REGION Network 21: FC_CARGA_RECETA
   RUNG wire#powerrail
      Contact( "flanco"."pHMI.Pls_CargarReceta" )
      "FC_CARGA_RECETA"("NRO RECETA" := "DB_Animación".Nro_Receta_Edición)
   END_RUNG
   // the same network as SCL:
   IF "flanco"."pHMI.Pls_CargarReceta" THEN
       "FC_CARGA_RECETA"("NRO RECETA" := "DB_Animación".Nro_Receta_Edición);
   END_IF;
END_REGION

REGION Network 22: Proceso a Animación
   RUNG wire#powerrail
      I_Contact( "Editando_Recetas" )
      "CAPA Proceso_Animación"()
   END_RUNG
   // the same network as SCL:
   IF NOT "Editando_Recetas" THEN "CAPA Proceso_Animación"(); END_IF;
END_REGION

REGION Network 23: CAPA Receta_Animación_Receta
   RUNG wire#powerrail
      "CAPA Receta_Animación_Receta"()
   END_RUNG
   // the same network as SCL:
   "CAPA Receta_Animación_Receta"();
END_REGION

REGION Network 24: Animación
   RUNG wire#powerrail
      "FC_Animación"()
   END_RUNG
   // the same network as SCL:
   "FC_Animación"();
END_REGION

REGION Network 25: RESET ELEM ACTUAL
   RUNG wire#powerrail
      I_Contact( "AUTO/MAN" )
      "FC_RESET_ELEM_ACTUAL"()
   END_RUNG
   // the same network as SCL:
   IF NOT "AUTO/MAN" THEN "FC_RESET_ELEM_ACTUAL"(); END_IF;
END_REGION

REGION Network 26: Alarmas
   RUNG wire#powerrail
      "10_FC_Alarmas"()
   END_RUNG
   // the same network as SCL:
   "10_FC_Alarmas"();
END_REGION

REGION Network 27: Salidas
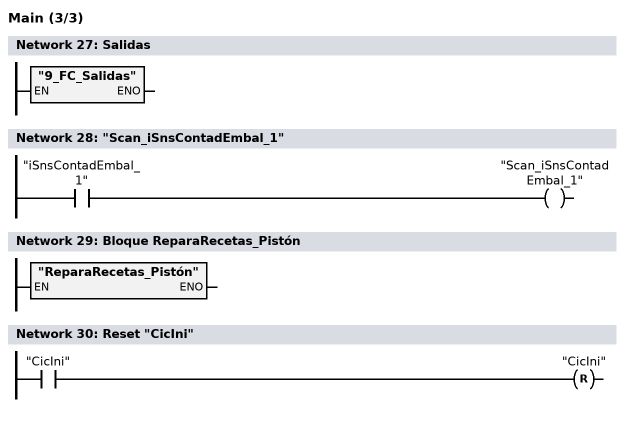
   RUNG wire#powerrail
      "9_FC_Salidas"()
   END_RUNG
   // the same network as SCL:
   "9_FC_Salidas"();
END_REGION

REGION Network 28: "Scan_iSnsContadEmbal_1"
   RUNG wire#powerrail
      Contact( "iSnsContadEmbal_1" )
      Coil( "Scan_iSnsContadEmbal_1" )
   END_RUNG
   // the same network as SCL:
   "Scan_iSnsContadEmbal_1" := "iSnsContadEmbal_1";
END_REGION

REGION Network 29: Bloque ReparaRecetas_Pistón
   RUNG wire#powerrail
      "ReparaRecetas_Pistón"()
   END_RUNG
   // the same network as SCL:
   "ReparaRecetas_Pistón"();
END_REGION

REGION Network 30: Reset "CicIni"
   RUNG wire#powerrail
      Contact( "CicIni" )
      R_Coil( "CicIni" )
   END_RUNG
   // the same network as SCL:
   IF "CicIni" THEN "CicIni" := FALSE; END_IF;
END_REGION
END_ORGANIZATION_BLOCK

ORGANIZATION_BLOCK "CYCL_FLT"   // OB80, LAD
TITLE = "Cycle Time Fault"
{ S7_Optimized_Access := 'FALSE' }
VERSION : 0.1
BEGIN
END_ORGANIZATION_BLOCK

ORGANIZATION_BLOCK "I/O_FLT1"   // OB82, LAD
TITLE = "I/O Point Fault"
{ S7_Optimized_Access := 'FALSE' }
VERSION : 0.1
BEGIN
END_ORGANIZATION_BLOCK

ORGANIZATION_BLOCK "OBNL_FLT"   // OB85, LAD
TITLE = "Organization Block (OB) Not Loaded Fault"
{ S7_Optimized_Access := 'FALSE' }
VERSION : 0.1
BEGIN
END_ORGANIZATION_BLOCK

ORGANIZATION_BLOCK "COMM_FLT"   // OB87, LAD
TITLE = "Communication Fault"
{ S7_Optimized_Access := 'FALSE' }
VERSION : 0.1
BEGIN
END_ORGANIZATION_BLOCK

ORGANIZATION_BLOCK "COMPLETE RESTART"   // OB100, LAD
TITLE = "Complete Restart"
{ S7_Optimized_Access := 'FALSE' }
VERSION : 0.1
BEGIN

REGION Network 1: "bit1"
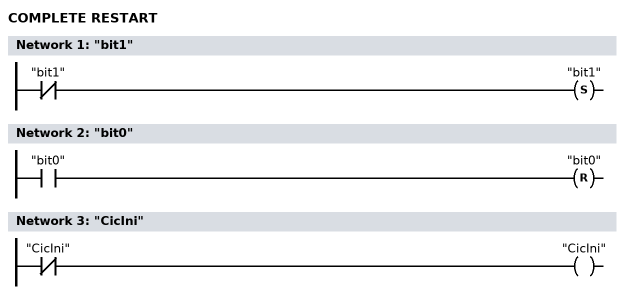
   RUNG wire#powerrail
      I_Contact( "bit1" )
      S_Coil( "bit1" )
   END_RUNG
   // the same network as SCL:
   IF NOT "bit1" THEN "bit1" := TRUE; END_IF;
END_REGION

REGION Network 2: "bit0"
   RUNG wire#powerrail
      Contact( "bit0" )
      R_Coil( "bit0" )
   END_RUNG
   // the same network as SCL:
   IF "bit0" THEN "bit0" := FALSE; END_IF;
END_REGION

REGION Network 3: "CicIni"
   RUNG wire#powerrail
      I_Contact( "CicIni" )
      Coil( "CicIni" )
   END_RUNG
   // the same network as SCL:
   "CicIni" := NOT "CicIni";
END_REGION
END_ORGANIZATION_BLOCK

ORGANIZATION_BLOCK "PROG_ERR"   // OB121, LAD
TITLE = "Programming Error"
{ S7_Optimized_Access := 'FALSE' }
VERSION : 0.1
BEGIN
END_ORGANIZATION_BLOCK

ORGANIZATION_BLOCK "MOD_ERR"   // OB122, LAD
TITLE = "Module Access Error"
{ S7_Optimized_Access := 'FALSE' }
VERSION : 0.1
BEGIN
END_ORGANIZATION_BLOCK

// folder: Alarmas

FUNCTION "10_FC_Alarmas" : Void   // FC23, LAD
{ S7_Optimized_Access := 'FALSE' }
VERSION : 0.1
BEGIN

REGION Network 1: Falla 1: Emergencia Almacén Pallets
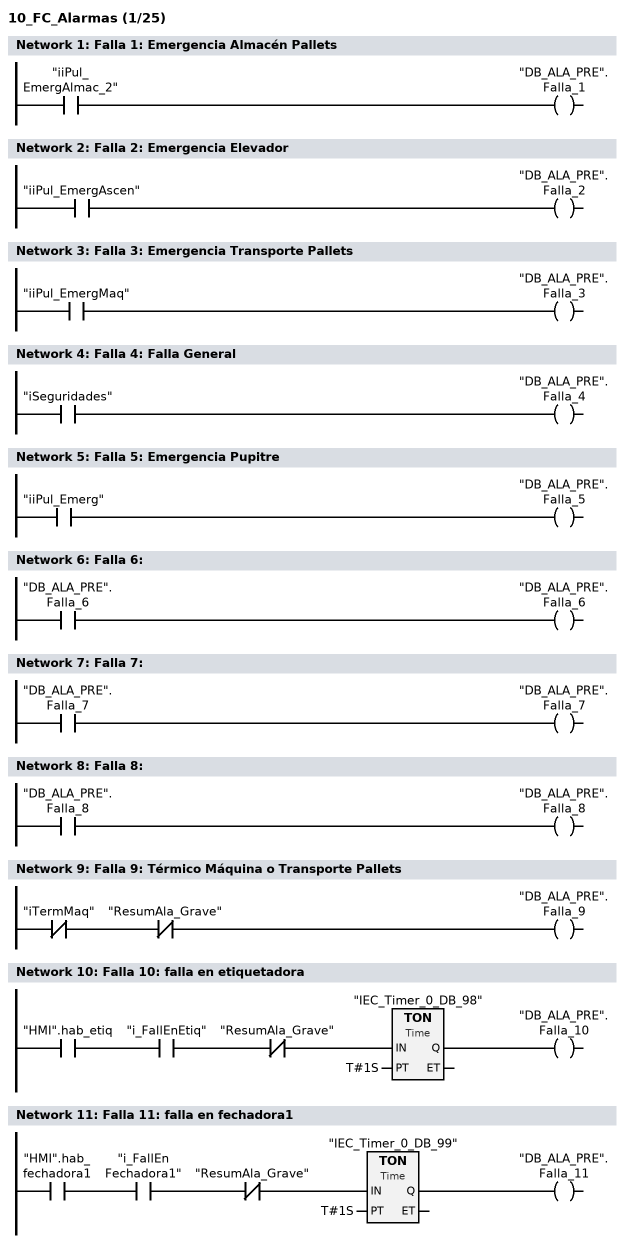
   RUNG wire#powerrail
      Contact( "iiPul_EmergAlmac_2" )
      Coil( "DB_ALA_PRE".Falla_1 )
   END_RUNG
   // the same network as SCL:
   "DB_ALA_PRE".Falla_1 := "iiPul_EmergAlmac_2";
END_REGION

REGION Network 2: Falla 2: Emergencia Elevador
   RUNG wire#powerrail
      Contact( "iiPul_EmergAscen" )
      Coil( "DB_ALA_PRE".Falla_2 )
   END_RUNG
   // the same network as SCL:
   "DB_ALA_PRE".Falla_2 := "iiPul_EmergAscen";
END_REGION

REGION Network 3: Falla 3: Emergencia Transporte Pallets
   RUNG wire#powerrail
      Contact( "iiPul_EmergMaq" )
      Coil( "DB_ALA_PRE".Falla_3 )
   END_RUNG
   // the same network as SCL:
   "DB_ALA_PRE".Falla_3 := "iiPul_EmergMaq";
END_REGION

REGION Network 4: Falla 4: Falla General
   RUNG wire#powerrail
      Contact( "iSeguridades" )
      Coil( "DB_ALA_PRE".Falla_4 )
   END_RUNG
   // the same network as SCL:
   "DB_ALA_PRE".Falla_4 := "iSeguridades";
END_REGION

REGION Network 5: Falla 5: Emergencia Pupitre
   RUNG wire#powerrail
      Contact( "iiPul_Emerg" )
      Coil( "DB_ALA_PRE".Falla_5 )
   END_RUNG
   // the same network as SCL:
   "DB_ALA_PRE".Falla_5 := "iiPul_Emerg";
END_REGION

REGION Network 6: Falla 6:
   RUNG wire#powerrail
      Contact( "DB_ALA_PRE".Falla_6 )
      Coil( "DB_ALA_PRE".Falla_6 )
   END_RUNG
   // the same network as SCL:
   "DB_ALA_PRE".Falla_6 := "DB_ALA_PRE".Falla_6;
END_REGION

REGION Network 7: Falla 7:
   RUNG wire#powerrail
      Contact( "DB_ALA_PRE".Falla_7 )
      Coil( "DB_ALA_PRE".Falla_7 )
   END_RUNG
   // the same network as SCL:
   "DB_ALA_PRE".Falla_7 := "DB_ALA_PRE".Falla_7;
END_REGION

REGION Network 8: Falla 8:
   RUNG wire#powerrail
      Contact( "DB_ALA_PRE".Falla_8 )
      Coil( "DB_ALA_PRE".Falla_8 )
   END_RUNG
   // the same network as SCL:
   "DB_ALA_PRE".Falla_8 := "DB_ALA_PRE".Falla_8;
END_REGION

REGION Network 9: Falla 9: Térmico Máquina o Transporte Pallets
   RUNG wire#powerrail
      I_Contact( "iTermMaq" )
      I_Contact( "ResumAla_Grave" )
      Coil( "DB_ALA_PRE".Falla_9 )
   END_RUNG
   // the same network as SCL:
   "DB_ALA_PRE".Falla_9 := NOT "iTermMaq" AND NOT "ResumAla_Grave";
END_REGION

REGION Network 10: Falla 10: falla en etiquetadora
   "IEC_Timer_0_DB_98".TON(IN := "HMI".hab_etiq AND "i_FallEnEtiq" AND NOT "ResumAla_Grave", PT := T#1S);
   "DB_ALA_PRE".Falla_10 := "IEC_Timer_0_DB_98".Q;
END_REGION

REGION Network 11: Falla 11: falla en fechadora1
   "IEC_Timer_0_DB_99".TON(IN := "HMI".hab_fechadora1 AND "i_FallEnFechadora1" AND NOT "ResumAla_Grave",
                           PT := T#1S);
   "DB_ALA_PRE".Falla_11 := "IEC_Timer_0_DB_99".Q;
END_REGION

REGION Network 12: Falla 12: falla en fechadora2
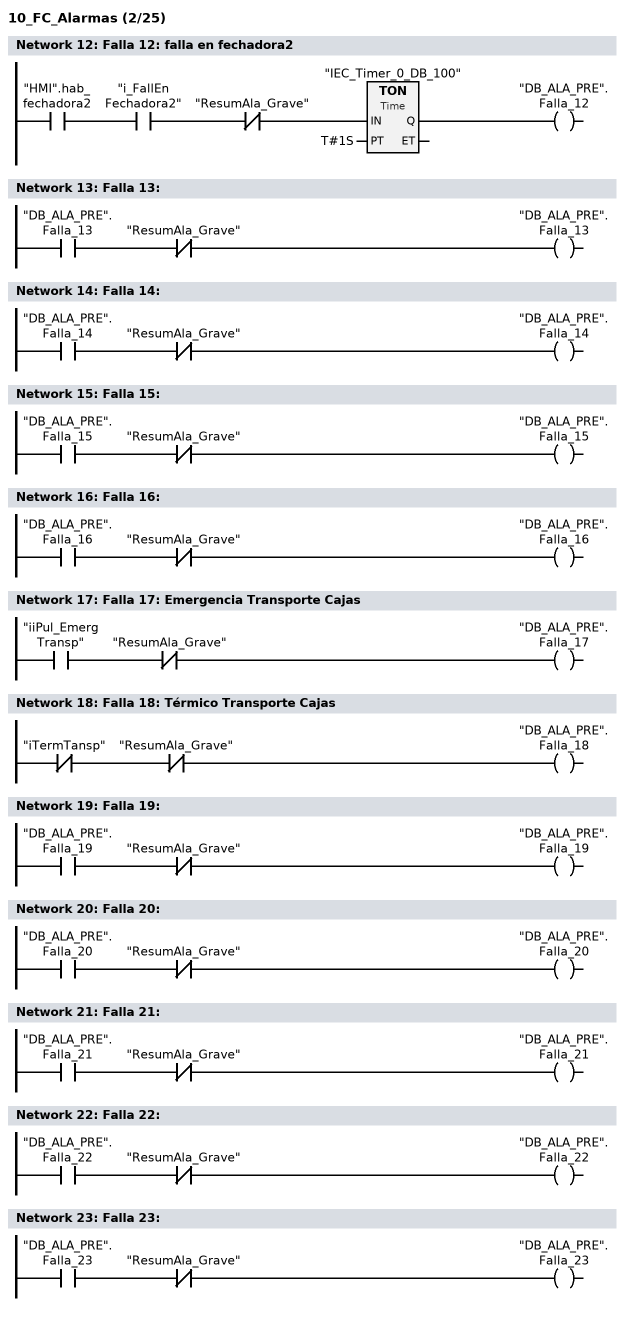
   "IEC_Timer_0_DB_100".TON(IN := "HMI".hab_fechadora2 AND "i_FallEnFechadora2" AND NOT "ResumAla_Grave",
                           PT := T#1S);
   "DB_ALA_PRE".Falla_12 := "IEC_Timer_0_DB_100".Q;
END_REGION

REGION Network 13: Falla 13:
   RUNG wire#powerrail
      Contact( "DB_ALA_PRE".Falla_13 )
      I_Contact( "ResumAla_Grave" )
      Coil( "DB_ALA_PRE".Falla_13 )
   END_RUNG
   // the same network as SCL:
   "DB_ALA_PRE".Falla_13 := "DB_ALA_PRE".Falla_13 AND NOT "ResumAla_Grave";
END_REGION

REGION Network 14: Falla 14:
   RUNG wire#powerrail
      Contact( "DB_ALA_PRE".Falla_14 )
      I_Contact( "ResumAla_Grave" )
      Coil( "DB_ALA_PRE".Falla_14 )
   END_RUNG
   // the same network as SCL:
   "DB_ALA_PRE".Falla_14 := "DB_ALA_PRE".Falla_14 AND NOT "ResumAla_Grave";
END_REGION

REGION Network 15: Falla 15:
   RUNG wire#powerrail
      Contact( "DB_ALA_PRE".Falla_15 )
      I_Contact( "ResumAla_Grave" )
      Coil( "DB_ALA_PRE".Falla_15 )
   END_RUNG
   // the same network as SCL:
   "DB_ALA_PRE".Falla_15 := "DB_ALA_PRE".Falla_15 AND NOT "ResumAla_Grave";
END_REGION

REGION Network 16: Falla 16:
   RUNG wire#powerrail
      Contact( "DB_ALA_PRE".Falla_16 )
      I_Contact( "ResumAla_Grave" )
      Coil( "DB_ALA_PRE".Falla_16 )
   END_RUNG
   // the same network as SCL:
   "DB_ALA_PRE".Falla_16 := "DB_ALA_PRE".Falla_16 AND NOT "ResumAla_Grave";
END_REGION

REGION Network 17: Falla 17: Emergencia Transporte Cajas
   RUNG wire#powerrail
      Contact( "iiPul_EmergTransp" )
      I_Contact( "ResumAla_Grave" )
      Coil( "DB_ALA_PRE".Falla_17 )
   END_RUNG
   // the same network as SCL:
   "DB_ALA_PRE".Falla_17 := "iiPul_EmergTransp" AND NOT "ResumAla_Grave";
END_REGION

REGION Network 18: Falla 18: Térmico Transporte Cajas
   RUNG wire#powerrail
      I_Contact( "iTermTansp" )
      I_Contact( "ResumAla_Grave" )
      Coil( "DB_ALA_PRE".Falla_18 )
   END_RUNG
   // the same network as SCL:
   "DB_ALA_PRE".Falla_18 := NOT "iTermTansp" AND NOT "ResumAla_Grave";
END_REGION

REGION Network 19: Falla 19:
   RUNG wire#powerrail
      Contact( "DB_ALA_PRE".Falla_19 )
      I_Contact( "ResumAla_Grave" )
      Coil( "DB_ALA_PRE".Falla_19 )
   END_RUNG
   // the same network as SCL:
   "DB_ALA_PRE".Falla_19 := "DB_ALA_PRE".Falla_19 AND NOT "ResumAla_Grave";
END_REGION

REGION Network 20: Falla 20:
   RUNG wire#powerrail
      Contact( "DB_ALA_PRE".Falla_20 )
      I_Contact( "ResumAla_Grave" )
      Coil( "DB_ALA_PRE".Falla_20 )
   END_RUNG
   // the same network as SCL:
   "DB_ALA_PRE".Falla_20 := "DB_ALA_PRE".Falla_20 AND NOT "ResumAla_Grave";
END_REGION

REGION Network 21: Falla 21:
   RUNG wire#powerrail
      Contact( "DB_ALA_PRE".Falla_21 )
      I_Contact( "ResumAla_Grave" )
      Coil( "DB_ALA_PRE".Falla_21 )
   END_RUNG
   // the same network as SCL:
   "DB_ALA_PRE".Falla_21 := "DB_ALA_PRE".Falla_21 AND NOT "ResumAla_Grave";
END_REGION

REGION Network 22: Falla 22:
   RUNG wire#powerrail
      Contact( "DB_ALA_PRE".Falla_22 )
      I_Contact( "ResumAla_Grave" )
      Coil( "DB_ALA_PRE".Falla_22 )
   END_RUNG
   // the same network as SCL:
   "DB_ALA_PRE".Falla_22 := "DB_ALA_PRE".Falla_22 AND NOT "ResumAla_Grave";
END_REGION

REGION Network 23: Falla 23:
   RUNG wire#powerrail
      Contact( "DB_ALA_PRE".Falla_23 )
      I_Contact( "ResumAla_Grave" )
      Coil( "DB_ALA_PRE".Falla_23 )
   END_RUNG
   // the same network as SCL:
   "DB_ALA_PRE".Falla_23 := "DB_ALA_PRE".Falla_23 AND NOT "ResumAla_Grave";
END_REGION

REGION Network 24: Falla 24:
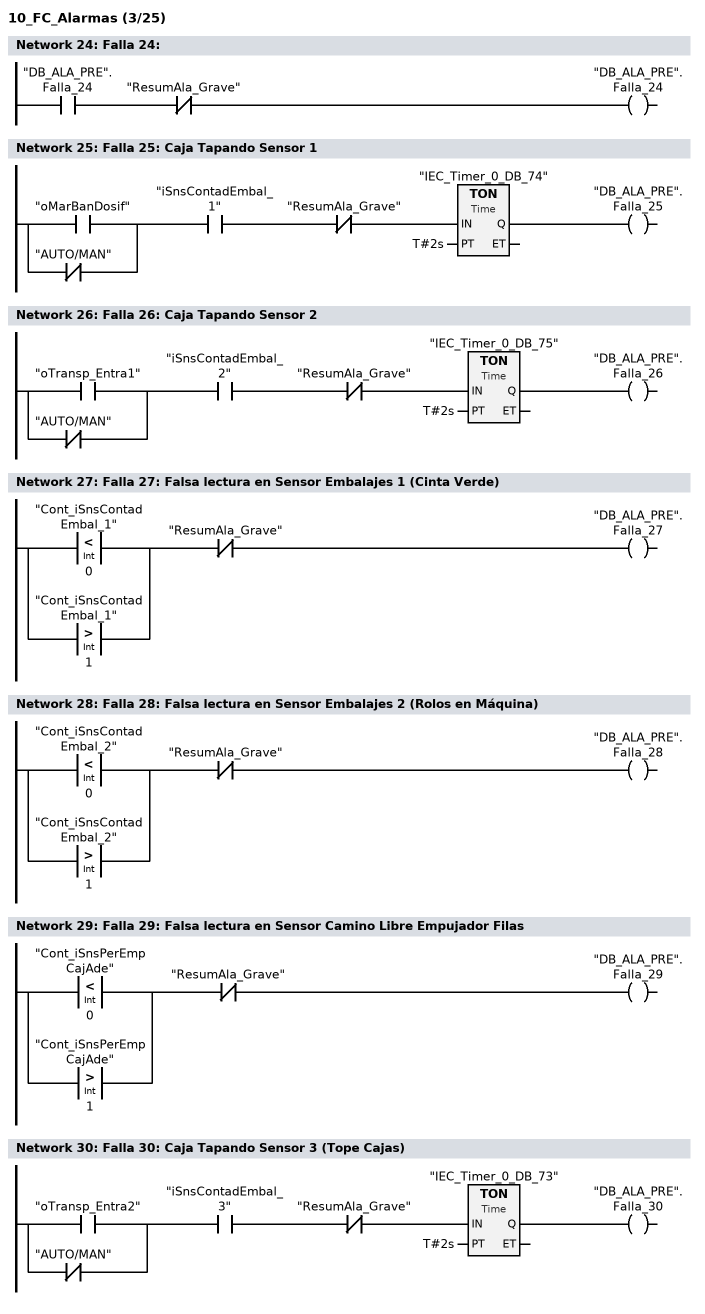
   RUNG wire#powerrail
      Contact( "DB_ALA_PRE".Falla_24 )
      I_Contact( "ResumAla_Grave" )
      Coil( "DB_ALA_PRE".Falla_24 )
   END_RUNG
   // the same network as SCL:
   "DB_ALA_PRE".Falla_24 := "DB_ALA_PRE".Falla_24 AND NOT "ResumAla_Grave";
END_REGION

REGION Network 25: Falla 25: Caja Tapando Sensor 1
   "IEC_Timer_0_DB_74".TON(IN := ("oMarBanDosif" OR NOT "AUTO/MAN") AND "iSnsContadEmbal_1" AND NOT "ResumAla_Grave",
                           PT := T#2s);
   "DB_ALA_PRE".Falla_25 := "IEC_Timer_0_DB_74".Q;
END_REGION

REGION Network 26: Falla 26: Caja Tapando Sensor 2
   "IEC_Timer_0_DB_75".TON(IN := ("oTransp_Entra1" OR NOT "AUTO/MAN") AND "iSnsContadEmbal_2" AND NOT "ResumAla_Grave",
                           PT := T#2s);
   "DB_ALA_PRE".Falla_26 := "IEC_Timer_0_DB_75".Q;
END_REGION

REGION Network 27: Falla 27: Falsa lectura en Sensor Embalajes 1 (Cinta Verde)
   RUNG wire#powerrail
      { S7_Templates := "SrcType := Int" } LT_Contact(in1 := "Cont_iSnsContadEmbal_1", in2 := 0)
      wire#w1
      I_Contact( "ResumAla_Grave" )
      Coil( "DB_ALA_PRE".Falla_27 )
   END_RUNG
   RUNG wire#powerrail
      { S7_Templates := "SrcType := Int" } GT_Contact(in1 := "Cont_iSnsContadEmbal_1", in2 := 1)
   END_RUNG wire#w1
   // the same network as SCL:
   "DB_ALA_PRE".Falla_27 := (("Cont_iSnsContadEmbal_1" < 0) OR ("Cont_iSnsContadEmbal_1" > 1)) AND NOT "ResumAla_Grave";
END_REGION

REGION Network 28: Falla 28: Falsa lectura en Sensor Embalajes 2 (Rolos en Máquina)
   RUNG wire#powerrail
      { S7_Templates := "SrcType := Int" } LT_Contact(in1 := "Cont_iSnsContadEmbal_2", in2 := 0)
      wire#w1
      I_Contact( "ResumAla_Grave" )
      Coil( "DB_ALA_PRE".Falla_28 )
   END_RUNG
   RUNG wire#powerrail
      { S7_Templates := "SrcType := Int" } GT_Contact(in1 := "Cont_iSnsContadEmbal_2", in2 := 1)
   END_RUNG wire#w1
   // the same network as SCL:
   "DB_ALA_PRE".Falla_28 := (("Cont_iSnsContadEmbal_2" < 0) OR ("Cont_iSnsContadEmbal_2" > 1)) AND NOT "ResumAla_Grave";
END_REGION

REGION Network 29: Falla 29: Falsa lectura en Sensor Camino Libre Empujador Filas
   RUNG wire#powerrail
      { S7_Templates := "SrcType := Int" } LT_Contact(in1 := "Cont_iSnsPerEmpCajAde", in2 := 0)
      wire#w1
      I_Contact( "ResumAla_Grave" )
      Coil( "DB_ALA_PRE".Falla_29 )
   END_RUNG
   RUNG wire#powerrail
      { S7_Templates := "SrcType := Int" } GT_Contact(in1 := "Cont_iSnsPerEmpCajAde", in2 := 1)
   END_RUNG wire#w1
   // the same network as SCL:
   "DB_ALA_PRE".Falla_29 := (("Cont_iSnsPerEmpCajAde" < 0) OR ("Cont_iSnsPerEmpCajAde" > 1)) AND NOT "ResumAla_Grave";
END_REGION

REGION Network 30: Falla 30: Caja Tapando Sensor 3 (Tope Cajas)
   "IEC_Timer_0_DB_73".TON(IN := ("oTransp_Entra2" OR NOT "AUTO/MAN") AND "iSnsContadEmbal_3" AND NOT "ResumAla_Grave",
                           PT := T#2s);
   "DB_ALA_PRE".Falla_30 := "IEC_Timer_0_DB_73".Q;
END_REGION

REGION Network 31: Falla 31: Falsa lectura en Sensor Embalajes 3 (Tope Cajas)
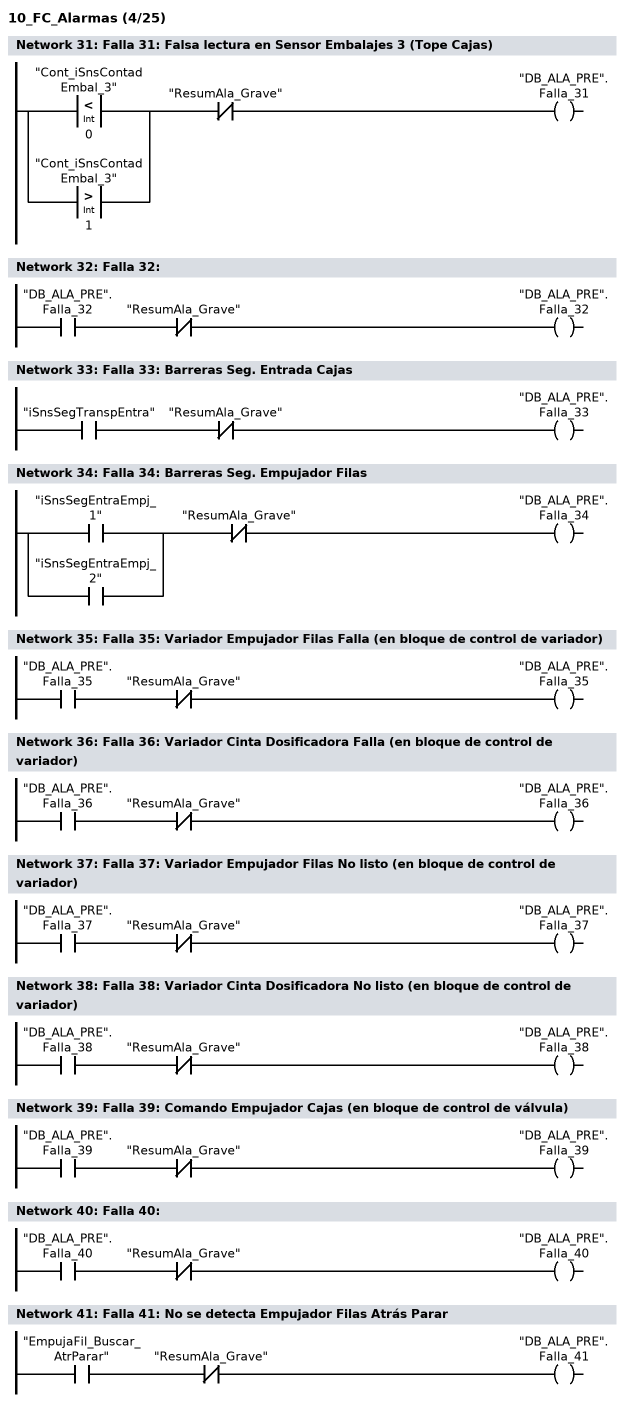
   RUNG wire#powerrail
      { S7_Templates := "SrcType := Int" } LT_Contact(in1 := "Cont_iSnsContadEmbal_3", in2 := 0)
      wire#w1
      I_Contact( "ResumAla_Grave" )
      Coil( "DB_ALA_PRE".Falla_31 )
   END_RUNG
   RUNG wire#powerrail
      { S7_Templates := "SrcType := Int" } GT_Contact(in1 := "Cont_iSnsContadEmbal_3", in2 := 1)
   END_RUNG wire#w1
   // the same network as SCL:
   "DB_ALA_PRE".Falla_31 := (("Cont_iSnsContadEmbal_3" < 0) OR ("Cont_iSnsContadEmbal_3" > 1)) AND NOT "ResumAla_Grave";
END_REGION

REGION Network 32: Falla 32:
   RUNG wire#powerrail
      Contact( "DB_ALA_PRE".Falla_32 )
      I_Contact( "ResumAla_Grave" )
      Coil( "DB_ALA_PRE".Falla_32 )
   END_RUNG
   // the same network as SCL:
   "DB_ALA_PRE".Falla_32 := "DB_ALA_PRE".Falla_32 AND NOT "ResumAla_Grave";
END_REGION

REGION Network 33: Falla 33: Barreras Seg. Entrada Cajas
   RUNG wire#powerrail
      Contact( "iSnsSegTranspEntra" )
      I_Contact( "ResumAla_Grave" )
      Coil( "DB_ALA_PRE".Falla_33 )
   END_RUNG
   // the same network as SCL:
   "DB_ALA_PRE".Falla_33 := "iSnsSegTranspEntra" AND NOT "ResumAla_Grave";
END_REGION

REGION Network 34: Falla 34: Barreras Seg. Empujador Filas
   RUNG wire#powerrail
      Contact( "iSnsSegEntraEmpj_1" )
      wire#w1
      I_Contact( "ResumAla_Grave" )
      Coil( "DB_ALA_PRE".Falla_34 )
   END_RUNG
   RUNG wire#powerrail
      Contact( "iSnsSegEntraEmpj_2" )
   END_RUNG wire#w1
   // the same network as SCL:
   "DB_ALA_PRE".Falla_34 := ("iSnsSegEntraEmpj_1" OR "iSnsSegEntraEmpj_2") AND NOT "ResumAla_Grave";
END_REGION

REGION Network 35: Falla 35: Variador Empujador Filas Falla (en bloque de control de variador)
   RUNG wire#powerrail
      Contact( "DB_ALA_PRE".Falla_35 )
      I_Contact( "ResumAla_Grave" )
      Coil( "DB_ALA_PRE".Falla_35 )
   END_RUNG
   // the same network as SCL:
   "DB_ALA_PRE".Falla_35 := "DB_ALA_PRE".Falla_35 AND NOT "ResumAla_Grave";
END_REGION

REGION Network 36: Falla 36: Variador Cinta Dosificadora Falla (en bloque de control de variador)
   RUNG wire#powerrail
      Contact( "DB_ALA_PRE".Falla_36 )
      I_Contact( "ResumAla_Grave" )
      Coil( "DB_ALA_PRE".Falla_36 )
   END_RUNG
   // the same network as SCL:
   "DB_ALA_PRE".Falla_36 := "DB_ALA_PRE".Falla_36 AND NOT "ResumAla_Grave";
END_REGION

REGION Network 37: Falla 37: Variador Empujador Filas No listo (en bloque de control de variador)
   RUNG wire#powerrail
      Contact( "DB_ALA_PRE".Falla_37 )
      I_Contact( "ResumAla_Grave" )
      Coil( "DB_ALA_PRE".Falla_37 )
   END_RUNG
   // the same network as SCL:
   "DB_ALA_PRE".Falla_37 := "DB_ALA_PRE".Falla_37 AND NOT "ResumAla_Grave";
END_REGION

REGION Network 38: Falla 38: Variador Cinta Dosificadora No listo (en bloque de control de variador)
   RUNG wire#powerrail
      Contact( "DB_ALA_PRE".Falla_38 )
      I_Contact( "ResumAla_Grave" )
      Coil( "DB_ALA_PRE".Falla_38 )
   END_RUNG
   // the same network as SCL:
   "DB_ALA_PRE".Falla_38 := "DB_ALA_PRE".Falla_38 AND NOT "ResumAla_Grave";
END_REGION

REGION Network 39: Falla 39: Comando Empujador Cajas (en bloque de control de válvula)
   RUNG wire#powerrail
      Contact( "DB_ALA_PRE".Falla_39 )
      I_Contact( "ResumAla_Grave" )
      Coil( "DB_ALA_PRE".Falla_39 )
   END_RUNG
   // the same network as SCL:
   "DB_ALA_PRE".Falla_39 := "DB_ALA_PRE".Falla_39 AND NOT "ResumAla_Grave";
END_REGION

REGION Network 40: Falla 40:
   RUNG wire#powerrail
      Contact( "DB_ALA_PRE".Falla_40 )
      I_Contact( "ResumAla_Grave" )
      Coil( "DB_ALA_PRE".Falla_40 )
   END_RUNG
   // the same network as SCL:
   "DB_ALA_PRE".Falla_40 := "DB_ALA_PRE".Falla_40 AND NOT "ResumAla_Grave";
END_REGION

REGION Network 41: Falla 41: No se detecta Empujador Filas Atrás Parar
   RUNG wire#powerrail
      Contact( "EmpujaFil_Buscar_AtrParar" )
      I_Contact( "ResumAla_Grave" )
      Coil( "DB_ALA_PRE".Falla_41 )
   END_RUNG
   // the same network as SCL:
   "DB_ALA_PRE".Falla_41 := "EmpujaFil_Buscar_AtrParar" AND NOT "ResumAla_Grave";
END_REGION

REGION Network 42: Falla 42: No se detecta Empujador Filas Atrás Lento
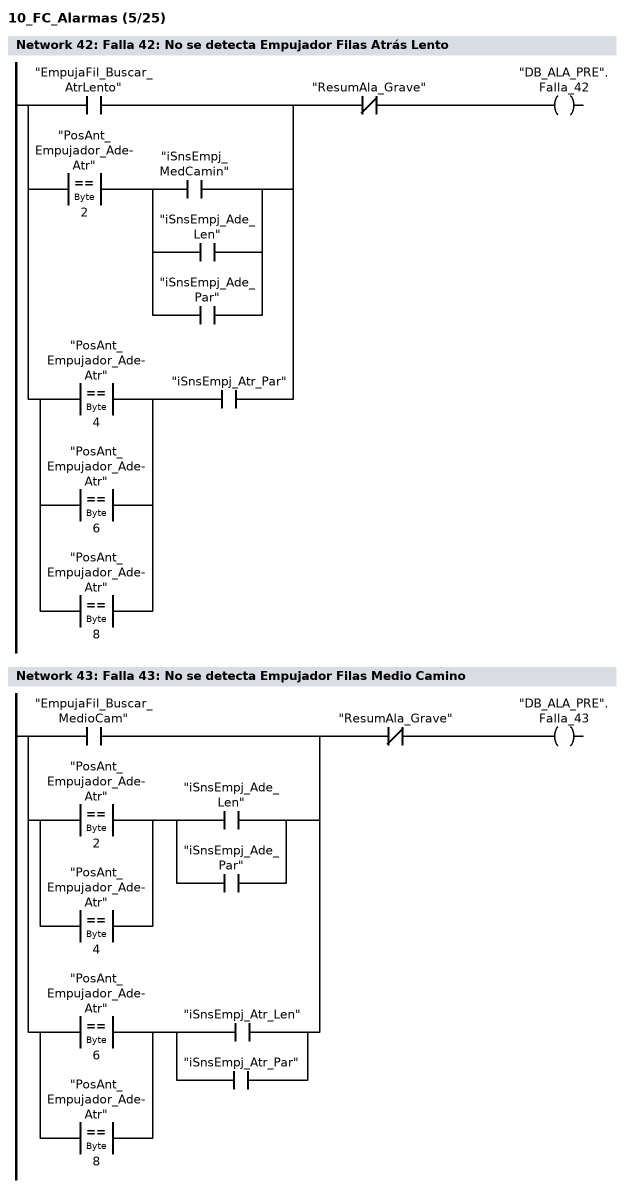
   RUNG wire#powerrail
      Contact( "EmpujaFil_Buscar_AtrLento" )
      wire#w1
      I_Contact( "ResumAla_Grave" )
      Coil( "DB_ALA_PRE".Falla_42 )
   END_RUNG
   RUNG wire#powerrail
      { S7_Templates := "SrcType := Byte" } EQ_Contact(in1 := "PosAnt_Empujador_Ade-Atr", in2 := 2)
      wire#w2
      Contact( "iSnsEmpj_MedCamin" )
   END_RUNG wire#w1
   RUNG wire#w2
      Contact( "iSnsEmpj_Ade_Len" )
   END_RUNG wire#w1
   RUNG wire#w2
      Contact( "iSnsEmpj_Ade_Par" )
   END_RUNG wire#w1
   RUNG wire#powerrail
      { S7_Templates := "SrcType := Byte" } EQ_Contact(in1 := "PosAnt_Empujador_Ade-Atr", in2 := 4)
      wire#w3
      Contact( "iSnsEmpj_Atr_Par" )
   END_RUNG wire#w1
   RUNG wire#powerrail
      { S7_Templates := "SrcType := Byte" } EQ_Contact(in1 := "PosAnt_Empujador_Ade-Atr", in2 := 6)
   END_RUNG wire#w3
   RUNG wire#powerrail
      { S7_Templates := "SrcType := Byte" } EQ_Contact(in1 := "PosAnt_Empujador_Ade-Atr", in2 := 8)
   END_RUNG wire#w3
   // the same network as SCL:
   "DB_ALA_PRE".Falla_42 := ("EmpujaFil_Buscar_AtrLento" OR (("PosAnt_Empujador_Ade-Atr" = 2) AND ("iSnsEmpj_MedCamin" OR "iSnsEmpj_Ade_Len" OR "iSnsEmpj_Ade_Par")) OR ((("PosAnt_Empujador_Ade-Atr" = 4) OR ("PosAnt_Empujador_Ade-Atr" = 6) OR ("PosAnt_Empujador_Ade-Atr" = 8)) AND "iSnsEmpj_Atr_Par")) AND NOT "ResumAla_Grave";
END_REGION

REGION Network 43: Falla 43: No se detecta Empujador Filas Medio Camino
   RUNG wire#powerrail
      Contact( "EmpujaFil_Buscar_MedioCam" )
      wire#w1
      I_Contact( "ResumAla_Grave" )
      Coil( "DB_ALA_PRE".Falla_43 )
   END_RUNG
   RUNG wire#powerrail
      { S7_Templates := "SrcType := Byte" } EQ_Contact(in1 := "PosAnt_Empujador_Ade-Atr", in2 := 2)
      wire#w2
      Contact( "iSnsEmpj_Ade_Len" )
   END_RUNG wire#w1
   RUNG wire#powerrail
      { S7_Templates := "SrcType := Byte" } EQ_Contact(in1 := "PosAnt_Empujador_Ade-Atr", in2 := 4)
   END_RUNG wire#w2
   RUNG wire#w2
      Contact( "iSnsEmpj_Ade_Par" )
   END_RUNG wire#w1
   RUNG wire#powerrail
      { S7_Templates := "SrcType := Byte" } EQ_Contact(in1 := "PosAnt_Empujador_Ade-Atr", in2 := 6)
      wire#w3
      Contact( "iSnsEmpj_Atr_Len" )
   END_RUNG wire#w1
   RUNG wire#powerrail
      { S7_Templates := "SrcType := Byte" } EQ_Contact(in1 := "PosAnt_Empujador_Ade-Atr", in2 := 8)
   END_RUNG wire#w3
   RUNG wire#w3
      Contact( "iSnsEmpj_Atr_Par" )
   END_RUNG wire#w1
   // the same network as SCL:
   "DB_ALA_PRE".Falla_43 := ("EmpujaFil_Buscar_MedioCam" OR ((("PosAnt_Empujador_Ade-Atr" = 2) OR ("PosAnt_Empujador_Ade-Atr" = 4)) AND ("iSnsEmpj_Ade_Len" OR "iSnsEmpj_Ade_Par")) OR ((("PosAnt_Empujador_Ade-Atr" = 6) OR ("PosAnt_Empujador_Ade-Atr" = 8)) AND ("iSnsEmpj_Atr_Len" OR "iSnsEmpj_Atr_Par"))) AND NOT "ResumAla_Grave";
END_REGION

REGION Network 44: Falla 44: No se detecta Empujador Filas Adelante Lento
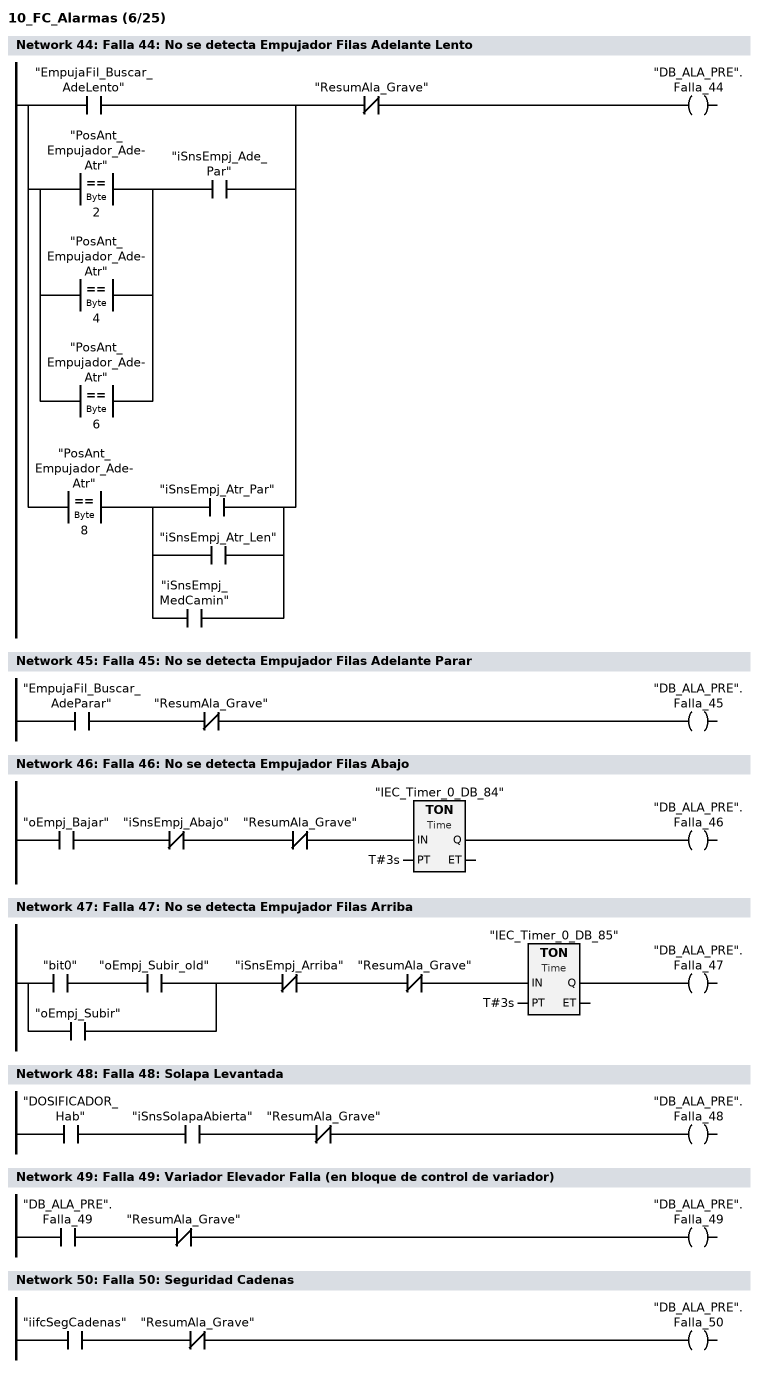
   RUNG wire#powerrail
      Contact( "EmpujaFil_Buscar_AdeLento" )
      wire#w1
      I_Contact( "ResumAla_Grave" )
      Coil( "DB_ALA_PRE".Falla_44 )
   END_RUNG
   RUNG wire#powerrail
      { S7_Templates := "SrcType := Byte" } EQ_Contact(in1 := "PosAnt_Empujador_Ade-Atr", in2 := 2)
      wire#w2
      Contact( "iSnsEmpj_Ade_Par" )
   END_RUNG wire#w1
   RUNG wire#powerrail
      { S7_Templates := "SrcType := Byte" } EQ_Contact(in1 := "PosAnt_Empujador_Ade-Atr", in2 := 4)
   END_RUNG wire#w2
   RUNG wire#powerrail
      { S7_Templates := "SrcType := Byte" } EQ_Contact(in1 := "PosAnt_Empujador_Ade-Atr", in2 := 6)
   END_RUNG wire#w2
   RUNG wire#powerrail
      { S7_Templates := "SrcType := Byte" } EQ_Contact(in1 := "PosAnt_Empujador_Ade-Atr", in2 := 8)
      wire#w3
      Contact( "iSnsEmpj_Atr_Par" )
   END_RUNG wire#w1
   RUNG wire#w3
      Contact( "iSnsEmpj_Atr_Len" )
   END_RUNG wire#w1
   RUNG wire#w3
      Contact( "iSnsEmpj_MedCamin" )
   END_RUNG wire#w1
   // the same network as SCL:
   "DB_ALA_PRE".Falla_44 := ("EmpujaFil_Buscar_AdeLento" OR ((("PosAnt_Empujador_Ade-Atr" = 2) OR ("PosAnt_Empujador_Ade-Atr" = 4) OR ("PosAnt_Empujador_Ade-Atr" = 6)) AND "iSnsEmpj_Ade_Par") OR (("PosAnt_Empujador_Ade-Atr" = 8) AND ("iSnsEmpj_Atr_Par" OR "iSnsEmpj_Atr_Len" OR "iSnsEmpj_MedCamin"))) AND NOT "ResumAla_Grave";
END_REGION

REGION Network 45: Falla 45: No se detecta Empujador Filas Adelante Parar
   RUNG wire#powerrail
      Contact( "EmpujaFil_Buscar_AdeParar" )
      I_Contact( "ResumAla_Grave" )
      Coil( "DB_ALA_PRE".Falla_45 )
   END_RUNG
   // the same network as SCL:
   "DB_ALA_PRE".Falla_45 := "EmpujaFil_Buscar_AdeParar" AND NOT "ResumAla_Grave";
END_REGION

REGION Network 46: Falla 46: No se detecta Empujador Filas Abajo
   "IEC_Timer_0_DB_84".TON(IN := "oEmpj_Bajar" AND NOT "iSnsEmpj_Abajo" AND NOT "ResumAla_Grave", PT := T#3s);
   "DB_ALA_PRE".Falla_46 := "IEC_Timer_0_DB_84".Q;
END_REGION

REGION Network 47: Falla 47: No se detecta Empujador Filas Arriba
   "IEC_Timer_0_DB_85".TON(IN := (("bit0" AND "oEmpj_Subir_old") OR "oEmpj_Subir") AND NOT "iSnsEmpj_Arriba" AND NOT "ResumAla_Grave",
                           PT := T#3s);
   "DB_ALA_PRE".Falla_47 := "IEC_Timer_0_DB_85".Q;
END_REGION

REGION Network 48: Falla 48: Solapa Levantada
   RUNG wire#powerrail
      Contact( "DOSIFICADOR_Hab" )
      Contact( "iSnsSolapaAbierta" )
      I_Contact( "ResumAla_Grave" )
      Coil( "DB_ALA_PRE".Falla_48 )
   END_RUNG
   // the same network as SCL:
   "DB_ALA_PRE".Falla_48 := "DOSIFICADOR_Hab" AND "iSnsSolapaAbierta" AND NOT "ResumAla_Grave";
END_REGION

REGION Network 49: Falla 49: Variador Elevador Falla (en bloque de control de variador)
   RUNG wire#powerrail
      Contact( "DB_ALA_PRE".Falla_49 )
      I_Contact( "ResumAla_Grave" )
      Coil( "DB_ALA_PRE".Falla_49 )
   END_RUNG
   // the same network as SCL:
   "DB_ALA_PRE".Falla_49 := "DB_ALA_PRE".Falla_49 AND NOT "ResumAla_Grave";
END_REGION

REGION Network 50: Falla 50: Seguridad Cadenas
   RUNG wire#powerrail
      Contact( "iifcSegCadenas" )
      I_Contact( "ResumAla_Grave" )
      Coil( "DB_ALA_PRE".Falla_50 )
   END_RUNG
   // the same network as SCL:
   "DB_ALA_PRE".Falla_50 := "iifcSegCadenas" AND NOT "ResumAla_Grave";
END_REGION

REGION Network 51: Falla 51: Seguridad Superior Elevador
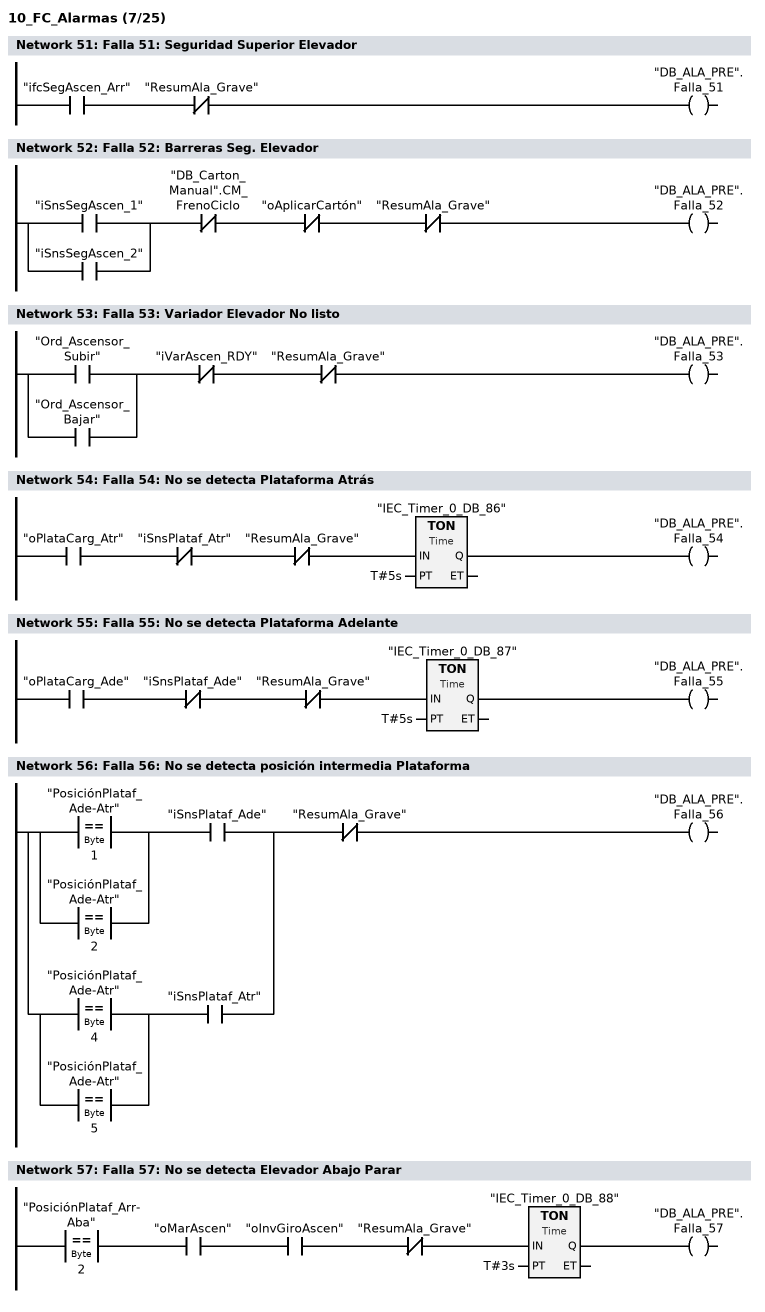
   RUNG wire#powerrail
      Contact( "ifcSegAscen_Arr" )
      I_Contact( "ResumAla_Grave" )
      Coil( "DB_ALA_PRE".Falla_51 )
   END_RUNG
   // the same network as SCL:
   "DB_ALA_PRE".Falla_51 := "ifcSegAscen_Arr" AND NOT "ResumAla_Grave";
END_REGION

REGION Network 52: Falla 52: Barreras Seg. Elevador
   RUNG wire#powerrail
      Contact( "iSnsSegAscen_1" )
      wire#w1
      I_Contact( "DB_Carton_Manual".CM_FrenoCiclo )
      I_Contact( "oAplicarCartón" )
      I_Contact( "ResumAla_Grave" )
      Coil( "DB_ALA_PRE".Falla_52 )
   END_RUNG
   RUNG wire#powerrail
      Contact( "iSnsSegAscen_2" )
   END_RUNG wire#w1
   // the same network as SCL:
   "DB_ALA_PRE".Falla_52 := ("iSnsSegAscen_1" OR "iSnsSegAscen_2") AND NOT "DB_Carton_Manual".CM_FrenoCiclo AND NOT "oAplicarCartón" AND NOT "ResumAla_Grave";
END_REGION

REGION Network 53: Falla 53: Variador Elevador No listo
   RUNG wire#powerrail
      Contact( "Ord_Ascensor_Subir" )
      wire#w1
      I_Contact( "iVarAscen_RDY" )
      I_Contact( "ResumAla_Grave" )
      Coil( "DB_ALA_PRE".Falla_53 )
   END_RUNG
   RUNG wire#powerrail
      Contact( "Ord_Ascensor_Bajar" )
   END_RUNG wire#w1
   // the same network as SCL:
   "DB_ALA_PRE".Falla_53 := ("Ord_Ascensor_Subir" OR "Ord_Ascensor_Bajar") AND NOT "iVarAscen_RDY" AND NOT "ResumAla_Grave";
END_REGION

REGION Network 54: Falla 54: No se detecta Plataforma Atrás
   "IEC_Timer_0_DB_86".TON(IN := "oPlataCarg_Atr" AND NOT "iSnsPlataf_Atr" AND NOT "ResumAla_Grave", PT := T#5s);
   "DB_ALA_PRE".Falla_54 := "IEC_Timer_0_DB_86".Q;
END_REGION

REGION Network 55: Falla 55: No se detecta Plataforma Adelante
   "IEC_Timer_0_DB_87".TON(IN := "oPlataCarg_Ade" AND NOT "iSnsPlataf_Ade" AND NOT "ResumAla_Grave", PT := T#5s);
   "DB_ALA_PRE".Falla_55 := "IEC_Timer_0_DB_87".Q;
END_REGION

REGION Network 56: Falla 56: No se detecta posición intermedia Plataforma
   RUNG wire#powerrail
      { S7_Templates := "SrcType := Byte" } EQ_Contact(in1 := "PosiciónPlataf_Ade-Atr", in2 := 1)
      wire#w1
      Contact( "iSnsPlataf_Ade" )
      wire#w2
      I_Contact( "ResumAla_Grave" )
      Coil( "DB_ALA_PRE".Falla_56 )
   END_RUNG
   RUNG wire#powerrail
      { S7_Templates := "SrcType := Byte" } EQ_Contact(in1 := "PosiciónPlataf_Ade-Atr", in2 := 2)
   END_RUNG wire#w1
   RUNG wire#powerrail
      { S7_Templates := "SrcType := Byte" } EQ_Contact(in1 := "PosiciónPlataf_Ade-Atr", in2 := 4)
      wire#w3
      Contact( "iSnsPlataf_Atr" )
   END_RUNG wire#w2
   RUNG wire#powerrail
      { S7_Templates := "SrcType := Byte" } EQ_Contact(in1 := "PosiciónPlataf_Ade-Atr", in2 := 5)
   END_RUNG wire#w3
   // the same network as SCL:
   "DB_ALA_PRE".Falla_56 := (((("PosiciónPlataf_Ade-Atr" = 1) OR ("PosiciónPlataf_Ade-Atr" = 2)) AND "iSnsPlataf_Ade") OR ((("PosiciónPlataf_Ade-Atr" = 4) OR ("PosiciónPlataf_Ade-Atr" = 5)) AND "iSnsPlataf_Atr")) AND NOT "ResumAla_Grave";
END_REGION

REGION Network 57: Falla 57: No se detecta Elevador Abajo Parar
   "IEC_Timer_0_DB_88".TON(IN := ("PosiciónPlataf_Arr-Aba" = 2) AND "oMarAscen" AND "oInvGiroAscen" AND NOT "ResumAla_Grave",
                           PT := T#3s);
   "DB_ALA_PRE".Falla_57 := "IEC_Timer_0_DB_88".Q;
END_REGION

REGION Network 58: Falla 58: No se detecta Elevador Abajo Lento
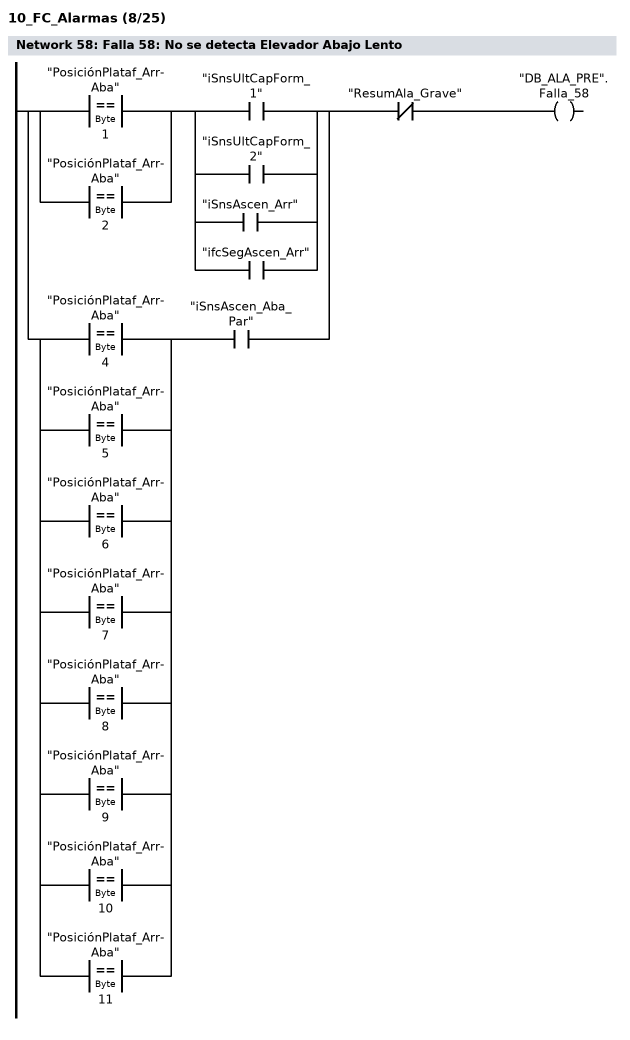
   RUNG wire#powerrail
      { S7_Templates := "SrcType := Byte" } EQ_Contact(in1 := "PosiciónPlataf_Arr-Aba", in2 := 1)
      wire#w1
      Contact( "iSnsUltCapForm_1" )
      wire#w2
      I_Contact( "ResumAla_Grave" )
      Coil( "DB_ALA_PRE".Falla_58 )
   END_RUNG
   RUNG wire#powerrail
      { S7_Templates := "SrcType := Byte" } EQ_Contact(in1 := "PosiciónPlataf_Arr-Aba", in2 := 2)
   END_RUNG wire#w1
   RUNG wire#w1
      Contact( "iSnsUltCapForm_2" )
   END_RUNG wire#w2
   RUNG wire#w1
      Contact( "iSnsAscen_Arr" )
   END_RUNG wire#w2
   RUNG wire#w1
      Contact( "ifcSegAscen_Arr" )
   END_RUNG wire#w2
   RUNG wire#powerrail
      { S7_Templates := "SrcType := Byte" } EQ_Contact(in1 := "PosiciónPlataf_Arr-Aba", in2 := 4)
      wire#w3
      Contact( "iSnsAscen_Aba_Par" )
   END_RUNG wire#w2
   RUNG wire#powerrail
      { S7_Templates := "SrcType := Byte" } EQ_Contact(in1 := "PosiciónPlataf_Arr-Aba", in2 := 5)
   END_RUNG wire#w3
   RUNG wire#powerrail
      { S7_Templates := "SrcType := Byte" } EQ_Contact(in1 := "PosiciónPlataf_Arr-Aba", in2 := 6)
   END_RUNG wire#w3
   RUNG wire#powerrail
      { S7_Templates := "SrcType := Byte" } EQ_Contact(in1 := "PosiciónPlataf_Arr-Aba", in2 := 7)
   END_RUNG wire#w3
   RUNG wire#powerrail
      { S7_Templates := "SrcType := Byte" } EQ_Contact(in1 := "PosiciónPlataf_Arr-Aba", in2 := 8)
   END_RUNG wire#w3
   RUNG wire#powerrail
      { S7_Templates := "SrcType := Byte" } EQ_Contact(in1 := "PosiciónPlataf_Arr-Aba", in2 := 9)
   END_RUNG wire#w3
   RUNG wire#powerrail
      { S7_Templates := "SrcType := Byte" } EQ_Contact(in1 := "PosiciónPlataf_Arr-Aba", in2 := 10)
   END_RUNG wire#w3
   RUNG wire#powerrail
      { S7_Templates := "SrcType := Byte" } EQ_Contact(in1 := "PosiciónPlataf_Arr-Aba", in2 := 11)
   END_RUNG wire#w3
   // the same network as SCL:
   "DB_ALA_PRE".Falla_58 := (((("PosiciónPlataf_Arr-Aba" = 1) OR ("PosiciónPlataf_Arr-Aba" = 2)) AND ("iSnsUltCapForm_1" OR "iSnsUltCapForm_2" OR "iSnsAscen_Arr" OR "ifcSegAscen_Arr")) OR ((("PosiciónPlataf_Arr-Aba" = 4) OR ("PosiciónPlataf_Arr-Aba" = 5) OR ("PosiciónPlataf_Arr-Aba" = 6) OR ("PosiciónPlataf_Arr-Aba" = 7) OR ("PosiciónPlataf_Arr-Aba" = 8) OR ("PosiciónPlataf_Arr-Aba" = 9) OR ("PosiciónPlataf_Arr-Aba" = 10) OR ("PosiciónPlataf_Arr-Aba" = 11)) AND "iSnsAscen_Aba_Par")) AND NOT "ResumAla_Grave";
END_REGION

REGION Network 59: Falla 59: No se detecta
